VERSION : 1.0
   VAR_INPUT
      IN_iSourceIndex : Int;
      IN_iDestIndex : Int;
      IN_iCount : Int;
   END_VAR
   VAR_IN_OUT
      INO_vSourceArrayStruct : Variant;
      INO_vDestArrayStruct : Variant;
   END_VAR
BEGIN
   #GP_BlockMoveStruct :=  MOVE_BLK_VARIANT(SRC:=#INO_vSourceArrayStruct,
                                            COUNT:=INT_TO_UDINT(#IN_iCount),
                                            SRC_INDEX:=INT_TO_DINT(#IN_iSourceIndex),
                                            DEST_INDEX:=INT_TO_DINT(#IN_iDestIndex),
                                            DEST=>#INO_vDestArrayStruct);
END_FUNCTION

// folder: TaskErrors

ORGANIZATION_BLOCK "Time error interrupt"   // OB80, LAD, TimeErrorInterrupt
{ S7_Optimized_Access := 'TRUE' }
VERSION : 0.1
   VAR_INPUT
      Fault_ID : Byte;   // Fault identifier
      Csg_OBnr : OB_Any;   // Number of OB causing the error
      Csg_Prio : UInt;   // Priority of OB causing the error
   END_VAR
BEGIN
END_ORGANIZATION_BLOCK

ORGANIZATION_BLOCK "Diagnostic error interrupt"   // OB82, LAD, DiagnosticErrorInterrupt
{ S7_Optimized_Access := 'TRUE' }
VERSION : 0.1
   VAR_INPUT
      IO_State : Word;   // IO state of the HW object
      LADDR : Hw_Any;   // Hardware identifier
      Channel : UInt;   // Channel number
      MultiError : Bool;   // =true if more than one error is present
   END_VAR
   VAR_TEMP
      RALM : Struct
         AINFO : "AINFO_";
         TINFO : "TINFO_";
         RETVAL : Int;
         ALLARMI_da_OB82 : Struct
            RALM : "PN_Alarm";
            LADDR : Hw_Any;
            evento_uscente : Bool;
         END_STRUCT;
      END_STRUCT;
      TMP_dId : DInt;
   END_VAR
BEGIN

REGION Network 1
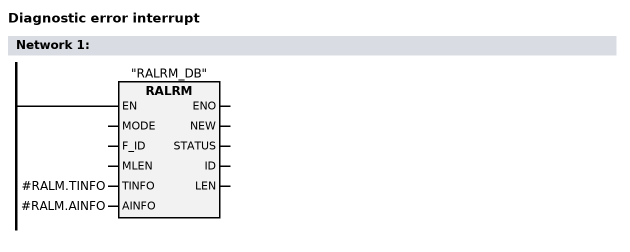
   "RALRM_DB"(TINFO := #RALM.TINFO, AINFO := #RALM.AINFO);   // RALRM
END_REGION

REGION Network 2 (SCL): Set alarms
   #TMP_dId:=UINT_TO_DINT("RALRM_DB".ID);

   IF "RALRM_DB".NEW THEN
       CASE #TMP_dId OF
           1:
               "RALRM_AUX_DB".tAlm.tF.xDevice1 := 1;
           2:
               "RALRM_AUX_DB".tAlm.tF.xDevice2 := 1;
           3:
               "RALRM_AUX_DB".tAlm.tF.xDevice3 := 1;
           4:
               "RALRM_AUX_DB".tAlm.tF.xDevice4 := 1;
           5:
               "RALRM_AUX_DB".tAlm.tF.xDevice5 := 1;
           6:
               "RALRM_AUX_DB".tAlm.tF.xDevice6 := 1;
           7:
               "RALRM_AUX_DB".tAlm.tF.xDevice7 := 1;
           8:
               "RALRM_AUX_DB".tAlm.tF.xDevice8 := 1;
           9:
               "RALRM_AUX_DB".tAlm.tF.xDevice9 := 1;
           10:
               "RALRM_AUX_DB".tAlm.tF.xDevice10 := 1;
           ELSE
               ;
       END_CASE;
   END_IF;
END_REGION
END_ORGANIZATION_BLOCK

ORGANIZATION_BLOCK "Pull or plug of modules"   // OB83, LAD, PullPlug
{ S7_Optimized_Access := 'TRUE' }
VERSION : 0.1
   VAR_INPUT
      LADDR : Hw_Io;   // Hardware identifier
      Event_Class : Byte;   // 16#38/39: module inserted, removed
      Fault_ID : Byte;   // Fault identifier
   END_VAR
BEGIN
END_ORGANIZATION_BLOCK

ORGANIZATION_BLOCK "Rack or station failure"   // OB86, LAD, RackStationFailure
{ S7_Optimized_Access := 'TRUE' }
VERSION : 0.1
   VAR_INPUT
      LADDR : Hw_Device;   // Hardware identifier
      Event_Class : Byte;   // Event class
      Fault_ID : Byte;   // Fault identifier
   END_VAR
BEGIN
END_ORGANIZATION_BLOCK

ORGANIZATION_BLOCK "Programming error"   // OB121, LAD, ProgrammingError
{ S7_Optimized_Access := 'TRUE' }
VERSION : 0.1
   VAR_INPUT
      BlockNr : UInt;   // Number of causing block
      Reaction : USInt;   // 0:ignore, 1:substitute, 2:skip
      Fault_ID : Byte;   // Fault identifier
      BlockType : USInt;   // 16#01:OB, 16#02:FC, 16#03:FB, 16#04:SFC, 16#05:SFB, 16#06:DB: Type of block causing the error
      Area : USInt;   // Area where the error occured
      DBNr : DB_ANY;   // DB number if Area = DB or DI
      Csg_OBNr : OB_Any;   // Number of OB causing the error
      Csg_Prio : USInt;   // Priority of OB causing the error
      Width : USInt;   // 0:bit, 1:byte, 2:word, 3:dword, 4:lword
   END_VAR
BEGIN
END_ORGANIZATION_BLOCK

ORGANIZATION_BLOCK "IO access error"   // OB122, LAD, IOAccessError
{ S7_Optimized_Access := 'TRUE' }
VERSION : 0.1
   VAR_INPUT
      BlockNr : UInt;   // Number of causing block
      Reaction : USInt;   // 0:ignore, 1:substitute, 2:skip
      Fault_ID : Byte;   // 16#42:reading, 16#43:writing
      BlockType : USInt;   // 16#01:OB, 16#02:FC, 16#03:FB, 16#04:SFC, 16#05:SFB, 16#06:DB: Type of block causing the error
      Area : USInt;   // 16#81:I, 16#82:Q: IO area where the IOaccess error occured
      DBNr : DB_ANY;   // Reserved for system
      Csg_OBNr : OB_Any;   // Number of OB causing the error
      Csg_Prio : USInt;   // Priority of OB causing the error
      Width : USInt;   // 0:bit, 1:byte, 2:word, 3:dword, 4:lword
   END_VAR
BEGIN
END_ORGANIZATION_BLOCK

// ===== PLC "1B160AP"  CPU 1512SP-1 PN =====

VAR_GLOBAL   // PLC tag table "Tabella delle variabili standard"
   "System_Byte" AT %MB0 : Byte;
   "FirstScan" AT %M0.0 : Bool;
   "DiagStatusUpdate" AT %M0.1 : Bool;
   "AlwaysTRUE" AT %M0.2 : Bool;
   "AlwaysFALSE" AT %M0.3 : Bool;
   "AlwaysOFF_Debug" AT %M10.0 : Bool;
   "o.1B160AP1.Open_SW_Gate" AT %Q39.0 : Bool;
   "i.1B160AP1.CounterActualValue" AT %ID30 : DWord;
   "i.1B160AP1.FrequencyActualValue" AT %ID38 : Real;
   "i.1B160AP1.CaptureValue" AT %ID34 : DWord;
   "o.1B160AP1.Res_Event" AT %Q40.1 : Bool;
   "o.1B160AP1.M217CutPressureHead1" AT %AW50 : Int;
   "o.1B160AP1.M217CutPressureHead2" AT %AW52 : Int;
   "o.1B160AP1.M217CutPressureHead5" AT %QW58 : Int;
   "o.1B160AP1.Enable_Measure" AT %Q39.7 : Bool;
   "i.1B160AP1.CounterCardStatus" AT %ED42 : DWord;
   "o.1B160AP1.CounterCardStatus" AT %AD38 : DWord;
   "o.1B160AP1.M217CutPressureHead3" AT %AW54 : Int;
   "o.1B160AP1.M217CutPressureHead4" AT %QW56 : Int;
   "o.IDeviceCPU0" AT %Q250.0 : "UDT_CM_IDEV_ToMainLine";
   "i.IDeviceCPU0" AT %I250.0 : "UDT_CM_IDEV_FromMainLine";
   "i.1B160AP1.Res_Event_Ack" AT %I43.1 : Bool;
   "i.1B160AP1.Event_Capture" AT %I45.6 : Bool;
   "cigliu" AT %M1.0 : Bool;
   "i.1B160AP1.1B18-2L+.PowerSupplyInputControlCabinetON" AT %E0.0 : Bool;
   "i.1B160AP1.1B18-3L+.InputInstallationPowerSupplyON" AT %E0.1 : Bool;
   "i.1B160AP1.1B11QF1/2.AnomalyPowerSupplies230V" AT %E0.2 : Bool;
   "i.1B160AP1.1B18QF2.PowerSupply24VLogic" AT %E0.3 : Bool;
   "i.1B160AP1.1B18QF3.PowerSupply24VLogic" AT %E0.4 : Bool;
   "i.1B160AP1.1B20QF2.PowerSupply24VLogic" AT %E0.5 : Bool;
   "i.1B160AP1.1B122KE1.MainEmergencyON" AT %E1.1 : Bool;
   "i.1B160AP1.1B41QF1.ProtectionPowerSupply36V_Motor_1-4" AT %I1.4 : Bool;
   "i.1B160AP1.1B41QF2.ProtectionPowerSupplyMotorsYcut_1-4" AT %I1.5 : Bool;
   "i.1B160AP1.1B51QM1.ProtectionCarriageTranslation" AT %E2.0 : Bool;
   "i.1B160AP1.1B52QM1.ProtectionCarriageTranslation" AT %E2.1 : Bool;
   "i.1B160AP1.1B53QM1.ProtectionCarriageTranslation" AT %E2.2 : Bool;
   "i.1B160AP1.1B54QM1.ProtectionCarriageTranslation" AT %E2.3 : Bool;
   "i.1B160AP1.1B55QM1.ProtectionCarriageTranslation" AT %I2.4 : Bool;
   "i.1B160AP1.M217B1SB1.LocalEmergency" AT %I3.1 : Bool;
   "i.1B160AP1.M217B1SB3_SB4.HeadsUpIstantaneous" AT %I3.0 : Bool;
   "i.1B411AP1.1B411SA1.Head1.CuttingPressure+" AT %E111.2 : Bool;
   "i.1B411AP1.1B411SQ1.Head1.CarriageHeadWorkPosition" AT %E111.3 : Bool;
   "i.1B411AP1.1B411SA1.Head1.CuttingPressure-" AT %E112.2 : Bool;
   "i.1B411AP1.1B411SA2.Head1.ProductionON" AT %E112.4 : Bool;
   "i.1B412AP1.1B412SA1.Head2.CuttingPressure+" AT %E121.2 : Bool;
   "i.1B412AP1.1B412SQ1.Head2.CarriageHeadWorkPosition" AT %E121.3 : Bool;
   "i.1B412AP1.1B412SA1.Head2.CuttingPressure-" AT %E122.2 : Bool;
   "i.1B412AP1.1B412SA2.Head2.ProductionON" AT %E122.4 : Bool;
   "i.1B413AP1.1B413SA1.Head3.CuttingPressure+" AT %E131.2 : Bool;
   "i.1B413AP1.1B413SQ1.Head3.CarriageHeadWorkPosition" AT %E131.3 : Bool;
   "i.1B413AP1.1B413SA1.Head3.CuttingPressure-" AT %E132.2 : Bool;
   "i.1B413AP1.1B413SA2.Head3.ProductionON" AT %E132.4 : Bool;
   "i.1B414AP1.1B414SA1.Head4.CuttingPressure+" AT %E141.2 : Bool;
   "i.1B414AP1.1B414SQ1.Head4.CarriageHeadWorkPosition" AT %E141.3 : Bool;
   "i.1B414AP1.1B414SA1.Head4.CuttingPressure-" AT %E142.2 : Bool;
   "i.1B414AP1.1B414SA2.Head4.ProductionON" AT %E142.4 : Bool;
   "i.1B415AP1.1B415SA1.Head5.CuttingPressure+" AT %I151.2 : Bool;
   "i.1B415AP1.1B415SQ1.Head5.CarriageHeadWorkPosition" AT %I151.3 : Bool;
   "i.1B415AP1.1B415SA1.Head5.CuttingPressure-" AT %I152.2 : Bool;
   "i.1B415AP1.1B415SA2.Head5.ProductionON" AT %I152.4 : Bool;
   "o.1B160AP1.1B251HL1.AreaFailure" AT %A0.0 : Bool;
   "o.1B160AP1.1B251KA1.ResetLocalEmergency" AT %A0.2 : Bool;
   "o.1B160AP1.EnableCard1" AT %A2.0 : Bool;
   "o.1B160AP1.EnableCard2" AT %A2.1 : Bool;
   "o.1B160AP1.EnableCard3" AT %A2.2 : Bool;
   "o.1B160AP1.EnableCard4" AT %A2.3 : Bool;
   "o.1B160AP1.EnableCard5" AT %Q2.4 : Bool;
   "o.1B160AP1.M217B1HL5.MachineToMaintenance" AT %Q0.6 : Bool;
   "o.1B160AP1.M217B1HL3.MachineReady" AT %Q0.4 : Bool;
   "o.1B160AP1.M217B1HL6.MachineOutOfOrder" AT %Q0.7 : Bool;
   "o.1B160AP1.M217B1HL4.MachineInOrder" AT %Q0.5 : Bool;
   "o.1B411AP1.1B411YV2.Head1.CuttingLubrication" AT %A111.0 : Bool;
   "o.1B411AP1.1B411YV1.Head1.CuttingHeadGlassApproach" AT %A111.1 : Bool;
   "o.1B411AP1.1B411SA2.Head1.ProductionON" AT %A111.4 : Bool;
   "o.1B412AP1.1B412YV2.Head2.CuttingLubrication" AT %A121.0 : Bool;
   "o.1B412AP1.1B412YV1.Head2.CuttingHeadGlassApproach" AT %A121.1 : Bool;
   "o.1B412AP1.1B412SA2.Head2.ProductionON" AT %A121.4 : Bool;
   "o.1B413AP1.1B413YV2.Head3.CuttingLubrication" AT %A131.0 : Bool;
   "o.1B413AP1.1B413YV1.Head3.CuttingHeadGlassApproach" AT %A131.1 : Bool;
   "o.1B413AP1.1B413SA2.Head3.ProductionON" AT %A131.4 : Bool;
   "o.1B414AP1.1B414YV2.Head4.CuttingLubrication" AT %A141.0 : Bool;
   "o.1B414AP1.1B414YV1.Head4.CuttingHeadGlassApproach" AT %A141.1 : Bool;
   "o.1B414AP1.1B414SA2.Head4.ProductionON" AT %A141.4 : Bool;
   "o.1B415AP1.1B415YV2.Head5.CuttingLubrication" AT %Q151.0 : Bool;
   "o.1B415AP1.1B415YV1.Head5.CuttingHeadGlassApproach" AT %Q151.1 : Bool;
   "o.1B415AP1.1B415SA2.Head5.ProductionON" AT %Q151.4 : Bool;
   "i.1B160AP1.1B20QF3.PowerSupply24VLogic" AT %I0.6 : Bool;
   "i.1B160AP1.1B42QF1.ProtectionPowerSupply36V_Motor_5-8" AT %I1.6 : Bool;
   "i.1B160AP1.1B42QF2.ProtectionPowerSupplyMotorsYcut_5-8" AT %I1.7 : Bool;
   "i.1B160AP1.1B56QM1.ProtectionCarriageTranslation" AT %I2.5 : Bool;
   "i.1B160AP1.1B57QM1.ProtectionCarriageTranslation" AT %I2.6 : Bool;
   "i.1B160AP1.1B58QM1.ProtectionCarriageTranslation" AT %I2.7 : Bool;
   "o.1B160AP1.EnableCard6" AT %Q2.5 : Bool;
   "o.1B160AP1.EnableCard7" AT %Q2.6 : Bool;
   "o.1B160AP1.EnableCard8" AT %Q2.7 : Bool;
   "o.1B160AP1.M217CutPressureHead6" AT %QW60 : Int;
   "o.1B160AP1.M217CutPressureHead7" AT %QW62 : Int;
   "o.1B160AP1.M217CutPressureHead8" AT %QW64 : Int;
   "o.1B416AP1.1B416SA2.Head6.ProductionON" AT %Q161.4 : Bool;
   "o.1B416AP1.1B416YV1.Head6.CuttingHeadGlassApproach" AT %Q161.1 : Bool;
   "o.1B416AP1.1B416YV2.Head6.CuttingLubrication" AT %Q161.0 : Bool;
   "o.1B417AP1.1B417SA2.Head7.ProductionON" AT %Q171.4 : Bool;
   "o.1B417AP1.1B417YV1.Head7.CuttingHeadGlassApproach" AT %Q171.1 : Bool;
   "o.1B417AP1.1B417YV2.Head7.CuttingLubrication" AT %Q171.0 : Bool;
   "o.1B418AP1.1B418SA2.Head8.ProductionON" AT %Q181.4 : Bool;
   "o.1B418AP1.1B418YV1.Head8.CuttingHeadGlassApproach" AT %Q181.1 : Bool;
   "o.1B418AP1.1B418YV2.Head8.CuttingLubrication" AT %Q181.0 : Bool;
   "i.1B416AP1.1B416SA1.Head6.CuttingPressure-" AT %I162.2 : Bool;
   "i.1B416AP1.1B416SA1.Head6.CuttingPressure+" AT %I161.2 : Bool;
   "i.1B416AP1.1B416SA2.Head6.ProductionON" AT %I162.4 : Bool;
   "i.1B416AP1.1B416SQ1.Head6.CarriageHeadWorkPosition" AT %I161.3 : Bool;
   "i.1B417AP1.1B417SA1.Head7.CuttingPressure-" AT %I172.2 : Bool;
   "i.1B417AP1.1B417SA1.Head7.CuttingPressure+" AT %I171.2 : Bool;
   "i.1B417AP1.1B417SA2.Head7.ProductionON" AT %I172.4 : Bool;
   "i.1B417AP1.1B417SQ1.Head7.CarriageHeadWorkPosition" AT %I171.3 : Bool;
   "i.1B418AP1.1B418SA1.Head8.CuttingPressure-" AT %I182.2 : Bool;
   "i.1B418AP1.1B418SA1.Head8.CuttingPressure+" AT %I181.2 : Bool;
   "i.1B418AP1.1B418SA2.Head8.ProductionON" AT %I182.4 : Bool;
   "i.1B418AP1.1B418SQ1.Head8.CarriageHeadWorkPosition" AT %I181.3 : Bool;
   "i.1B160AP1.M217B1SB2.LocalEmergency" AT %I3.2 : Bool;
END_VAR

VAR_GLOBAL CONSTANT   // PLC tag table "Tabella delle variabili standard"
   "CONST_dNumberOfHeadsCycle" : DInt := 7;   // Number of heads / Number of heads-1
   "CONST_dNumberOfHeads" : DInt := 8;   // Number of heads-1 / Number of heads
   "CONST_dPressureMax_MN" : DInt := 180000;   // Maximum allowable pressure [N/1000]
   "CONST_dPressureMin_MN" : DInt := 0;   // Minimum allowable pressure [N/1000]
   "CONST_dPressureMax_Unit" : DInt := 27648;   // Maximum allowable pressure Analog unit
   "CONST_dPressureMin_Unit" : DInt := 0;   // Minimum allowable pressure Analog unit
   "CONST_dFire_OnOff_MaxValue" : DInt := 5000;   // Fire ON OFF max value [mm/100]
   "CONST_dFire_OnOff_MinValue" : DInt := 0;   // Fire ON OFF min value [mm/100]
   "CONST_dPressureMax_Display_MN" : DInt := 180000;   // Maximum allowable pressure [N/1000]
   "CONST_dPressureMin_Display_MN" : DInt := 0;   // Minimum allowable pressure [N/1000]
   "CONST_dPressureMax_Display_Unit" : DInt := 27648;   // Maximum allowable pressure Analog unit
   "CONST_dPressureMin_Display_Unit" : DInt := 0;   // Minimum allowable pressure Analog unit
   "CONST_dPressureIncreasePneumatic_MN" : DInt := 250000;   // Pressure increse by cylinder [N/1000]
END_VAR

TYPE "ILx2T_Ref"
AUTHOR : SEMotion
FAMILY : LXM32
VERSION : 0.5
   STRUCT
      i_woDriveStatus : Word;
      i_by_ModeStatus : Byte;
      i_by_driveInput : Byte;
      i_wo_ActionWord : Word;
      i_wo_SpecialFunctions : Word;
      q_wo_dmControl : Word;
      q_dw_refA_16 : Word;
      q_dw_refB_32 : DWord;
      arOutputData : Array[0..7] of Byte;
      arInputData : Array[0..7] of Byte;
      stDriveStatus : Struct
         HaltActive : Bool;   // HALT is active
         reserved_Bit9 : Bool;
         reserved_Bit10 : Bool;
         reserved_Bit11 : Bool;
         reserved_Bit12 : Bool;
         x_Add : Bool;   // additional information
         x_End : Bool;   // OP mode finished - standstill
         x_Err : Bool;   // error
         state_Bit0 : Bool;   // Drive state bit 0
         state_Bit1 : Bool;   // Drive state bit 1
         state_Bit2 : Bool;   // Drive state bit 2
         state_Bit3 : Bool;   // Drive state bit 3
         reseverd_Bit4 : Bool;
         reserved_Bit5 : Bool;
         FaultActive : Bool;   // FAULT is active
         WarningActive : Bool;   // WARNING is active
      END_STRUCT;
      st_ModeStatus : Struct
         Mode_0 : Bool;   // Actual OP mode bit 0
         Mode_1 : Bool;   // Actual OP mode bit 1
         Mode_2 : Bool;   // Actual OP mode bit 2
         Mode_3 : Bool;   // Actual OP mode bit 3
         reserved : Bool;
         Reference_OK : Bool;   // drive is referenced
         ModeError : Bool;   // Status mode error
         ModeToggle : Bool;   // Status mode toggle
      END_STRUCT;
      st_ActionWord : Struct
         MotionNegative : Bool;   // negative direction
         InsidePosWindow : Bool;   // Inside Position Window
         reserved_Bit10 : Bool;
         TargetVelocityZero : Bool;   // Target velocity is zero
         Decelerating : Bool;
         Accelerating : Bool;
         ConstantVelocity : Bool;
         reserved_Bit15 : Bool;
         Reserved : Bool;
         Reserved_1 : Bool;
         Reserved_2 : Bool;
         Reserved_3 : Bool;
         Reserved_4 : Bool;
         Reserved_5 : Bool;
         MotionZero : Bool;   // Motion zero, actual velocity is zero
         MotionPositive : Bool;   // motor is moving in positiove direction
      END_STRUCT;
      st_SpecFunctions : Struct
         reserved_4 : Bool;   // Capture counter channel 1 bit 0
         reserved_5 : Bool;   // Capture counter channel 1 bit 1
         reserved_6 : Bool;   // Capture counter channel 2 bit 0
         reserved_7 : Bool;   // Capture counter channel 2 bit 1
         reserved_12 : Bool;
         reserved_13 : Bool;
         reserved_14 : Bool;
         reserved_15 : Bool;
         CAP1_0 : Bool;   // Actual OP mode bit 0
         CAP1_1 : Bool;   // Actual OP mode bit 1
         CAP2_0 : Bool;   // Actual OP mode bit 2
         CAP2_1 : Bool;   // Actual OP mode bit 3
         reserved : Bool;   // Actual OP mode bit 4
         reserved_1 : Bool;   // Status ModeDataError
         reserved_2 : Bool;   // Status mode error
         reserved_3 : Bool;   // Status mode toggle
      END_STRUCT;
      InitAccessID : Int;   // AccessID counter for INIT
      ProChAccessID : Int;   // Access ID Processchannel
      ParChAccessID : Int;   // Access ID Parameterchannel
      x_QuickStopInt : Bool;   // Library internal QuickStop Command
      x_FaultResetInt : Bool;   // Library internal FaultReset Command
      x_Set_HALT_Int : Bool;   // Library internal Set HALT Command
      x_Clear_HALT_Int : Bool;   // Library internal Clear HALT Command
      x_Continue_Int : Bool;   // Library internal HALT Contimue Command
      by_OP_ModeAct : Byte;   // Status - Actual operation mode
      x_IO_1 : Bool;   // Status of digital IO 1 (Bit 0)
      x_IO_2 : Bool;   // Status of digital IO 2 (Bit 1)
      x_IO_3 : Bool;   // Status of digital IO 3 (Bit 2)
      x_IO_4 : Bool;   // Status of digital IO 4 (Bit 3)
      x_STO_A : Bool;   // Status of Safe Torque Off Channel A
      x_STO_B : Bool;   // Status of Safe Torque Off Channel B
      x_reserved_6 : Bool;
      x_reserved_7 : Bool;
      x_CommandWriteParameter : Bool;
      x_CommandReadParameter : Bool;
      x_StatusReadParameter_OK : Bool;
      x_StatusReadParameter_Error : Bool;
      x_Status_WriteParameter_OK : Bool;
      x_Status_WriteParameter_Error : Bool;
      di_ParameterReadValue : DInt;
      di_ParameterWriteValue : DInt;
      udi_ModbusAddress_Read : UDInt;
      udi_ModbusAddress_Write : UDInt;
   END_STRUCT;
END_TYPE

TYPE "UDT_DataManager_HeadsBuffer"
VERSION : 0.1
   STRUCT
      rgdMissionID : Array[0..20] of DInt;   // Head#x mission ID
      rgdRequestPosition_cmm : Array[0..20] of DInt;   // Head#x request position [mm/100]
      rgdFireRequest : Array[0..20] of DInt;   // Head#x fire request
      dNumberOfElement : DInt;   // Number of element inside the buffer
   END_STRUCT;
END_TYPE

TYPE "UDT_DataManager_Insert"
VERSION : 0.1
   STRUCT
      dMissionCode : DInt;   // Mission code
      dMissionStart_cmm : DInt;   // Mission counter start [mm/100]
      dMissionEnd_cmm : DInt;   // Mission counter end [mm/100]
      rgxFireRequest : Array[0.."CONST_dNumberOfHeadsCycle"] of Bool;   // Fire request missions
      rgdHeadsPosition_cmm : Array[0.."CONST_dNumberOfHeadsCycle"] of DInt;   // Head#x position request [mm/100]
      xNewMission : Bool;   // New mission available
      xSystemReset : Bool;   // System reset
      rgdArmONReaction_ms : Array[0.."CONST_dNumberOfHeadsCycle"] of DInt;   // Head#x arm ON reaction [ms]
      rgdArmOFFReaction_ms : Array[0.."CONST_dNumberOfHeadsCycle"] of DInt;   // Head#x arm OFF reaction [ms]
      rgdFireONReaction_ms : Array[0.."CONST_dNumberOfHeadsCycle"] of DInt;   // Head#x fire ON reaction [ms]
      rgdFireOFFReaction_ms : Array[0.."CONST_dNumberOfHeadsCycle"] of DInt;   // Head#x fire OFF reaction [ms]
      rgdOilDelayStart_ms : Array[0.."CONST_dNumberOfHeadsCycle"] of DInt;   // Head#x oil delay start [ms]
      rgdOilDelayEnd_ms : Array[0.."CONST_dNumberOfHeadsCycle"] of DInt;   // Head#x oil advance end [ms]
      rgdFireONDelayStart_cmm : Array[0.."CONST_dNumberOfHeadsCycle"] of DInt;   // Head#x fire ON delay start [mm/100]
      rgdFireOFFDelayEnd_cmm : Array[0.."CONST_dNumberOfHeadsCycle"] of DInt;   // Head#x fire OFF delay end [mm/100]
   END_STRUCT;
END_TYPE

TYPE "UDT_DataManager"
VERSION : 0.1
   STRUCT
      tInputData : "UDT_DataManager_Insert";   // Manager input data
      tOutputData : "UDT_DataManager_Output";   // Manager output data
      dInterruptNumMissionTank : DInt;   // Number of mission fire inside the tank
      rgtInterruptMissionTank : Array[0..20] of "UDT_DataManager_Tank";   // Array of fire missions
      rgtOilList : Array[0.."CONST_dNumberOfHeadsCycle"] of "UDT_DataManager_HeadsBuffer";   // Oil list manager
      rgtArmList : Array[0.."CONST_dNumberOfHeadsCycle"] of "UDT_DataManager_HeadsBuffer";   // Arm list manager
   END_STRUCT;
END_TYPE

TYPE "UDT_DataManager_Output"
VERSION : 0.1
   STRUCT
      dMissionCode : DInt;   // Mission code number
      rgdFireHeadThreshold_cmm : Array[0.."CONST_dNumberOfHeadsCycle"] of DInt;   // Head#x firing threshold [mm/100]
      rgdHeadsPositions_cmm : Array[0.."CONST_dNumberOfHeadsCycle"] of DInt;   // Head#x positions request [mm/100]
      rgxFireHeadON_OFF : Array[0.."CONST_dNumberOfHeadsCycle"] of Bool;   // Head#x firing type request [bit]
      rgxDataToProcessInter : Array[0.."CONST_dNumberOfHeadsCycle"] of Bool;   // Head#x data to process by interrupt
      xGateOpen : Bool;   // Interrupt gate open
      dTargetLineValue_cmm : DInt;   // Virtual target line value [mm/100]
      rgxArmRequest : Array[0.."CONST_dNumberOfHeadsCycle"] of Bool;   // Head#x arming request
      rgdArmRequestTarget_cmm : Array[0.."CONST_dNumberOfHeadsCycle"] of DInt;   // Arm request target virtual [mm/100]
      rgxOilRequest : Array[0.."CONST_dNumberOfHeadsCycle"] of Bool;   // Head#x oil request
      rgdOilRequestTarget_cmm : Array[0.."CONST_dNumberOfHeadsCycle"] of DInt;   // Oil request target virtual [mm/100]
      rgdArmRequestIDMission : Array[0.."CONST_dNumberOfHeadsCycle"] of DInt;   // Arm request ID mission
      rgdOilRequestIDMission : Array[0.."CONST_dNumberOfHeadsCycle"] of DInt;   // Oil request ID mission
   END_STRUCT;
END_TYPE

TYPE "UDT_DataManager_Tank"
VERSION : 0.1
   STRUCT
      dMissionCode : DInt;   // Mission code
      dMissionValue_cmm : DInt;   // Mission value [mm/100]
      rgxFireRequest : Array[0.."CONST_dNumberOfHeadsCycle"] of Bool;   // Head#x fire request
      rgdHeadsPositions_cmm : Array[0.."CONST_dNumberOfHeadsCycle"] of DInt;   // Head#x position request [mm/100]
   END_STRUCT;
END_TYPE

TYPE "UDT_MB_ConnData"
   STRUCT
      IP_OCTET_1 : USInt;
      IP_OCTET_2 : USInt;
      IP_OCTET_3 : USInt;
      IP_OCTET_4 : USInt;
      ConnectID1 : Conn_Ouc;
      ConnectID2 : Conn_Ouc;
      ConnectID3 : Conn_Ouc;
      ConnectID4 : Conn_Ouc;
   END_STRUCT;
END_TYPE

TYPE "UDT_CM_IDEV_FromMainLine"
VERSION : 0.1
   STRUCT
      dSpare1 : Array[0..2] of DInt;
      xCycleON : Bool;   // Cycle ON
      xResetAnomaly : Bool;   // Reset anomaly
      xResetBuffers : Bool;   // Reset buffer
      xGlassBreak : Bool;   // Glass break under the bridge
      xPLCActive0 : Bool;   // PLC Active (0=CPU0, 1=CPU1)
      xPLCActive1 : Bool;   // PLC Active (0=CPU0, 1=CPU1)
      xQLTplate : Bool;   // Quality plate in progress
      xSpare2 : Bool;
      xSpare3 : Bool;
      xSpare4 : Bool;
      xSpare5 : Bool;
      xSpare6 : Bool;
      xSpare7 : Bool;
      xSpare8 : Bool;
      xSpare9 : Bool;
      xSpare10 : Bool;
      xStatusSpare : Array[0..15] of Bool;
      dSpare2 : Array[0..7] of DInt;
      iSpare : Int;
   END_STRUCT;
END_TYPE

TYPE "UDT_CM_IDEV_ToMainLine"
VERSION : 0.1
   STRUCT
      dProcessingIDPlate : DInt;   // Processing ID Plate [Num]
      dSpare1 : DInt;
      dSpare2 : DInt;
      rgxStatus : Array[0..31] of Bool;   // Status heads
      rgdHeadsPositions_cmm : Array[0..15] of DInt;   // Head #x position status
      rgxHeadStatus : Array[0..15] of Bool;   // Head #x enabled
      rgxCuttingStatus : Array[0..15] of Bool;   // Head #x cuuting status
      rgdHeadsPressure : Array[0..15] of DInt;   // Head #x Pressure [mN]
      rgrHeadsSpace : Array[0..15] of Real;   // Head #x Distance [Km]
      iFireOffset_ON : Int;   // All head fire on offset
      iFireOffset_OFF : Int;   // All head fire off offset
      iSpare : Int;
      dSpare : Array[0..7] of DInt;
   END_STRUCT;
   // // rgxStatus[0] : Glass break in progress
   // // rgxStatus[1] : Liftup pushbutton engaged
   // // rgxStatus[2] : Bridge enabled
   // // rgxStatus[3] : Bridge locked
   // // rgxStatus[8] : Fire offset calibration
END_TYPE

TYPE "UDT_CM_RECV_SyncroData"
VERSION : 0.1
   STRUCT
      dMissionID : DInt;   // Mission Identifier
      dSynchroValue_cmm : DInt;   // Counter value in the last synchro [mm/100]
      dSpare : Array[0..7] of DInt;
      xSpare : Array[0..15] of Bool;
      dSpare2 : Array[0..2] of DInt;
      iSpare : Int;
   END_STRUCT;
END_TYPE

TYPE "UDT_CM_RECV_MissionData"
VERSION : 0.1
   STRUCT
      dMissionID : DInt;   // Mission Identifier
      dMissionStart_cmm : DInt;   // Mission counter start [mm/100]
      dMissionEnd_cmm : DInt;   // Mission counter stop [mm/100]
      dTrackingDbNumber : DInt;   // Tracking DB number
      dSpare1 : Array[0..9] of DInt;
      rgxFireRequest : Array[0..31] of Bool;   // Head #x firing request
      rgdHeadsPosition_cmm : Array[0..15] of DInt;   // Head #x position request [mm/100]
      dSpare2 : Array[0..14] of DInt;
   END_STRUCT;
END_TYPE

TYPE "UDT_CM_Manager"
VERSION : 0.1
   STRUCT
      ST_xNewDataReceiveCPU0 : Bool;   // New data receive
      ST_xErrorCPU0 : Bool;   // Error
      ST_xNewSynchCPU0 : Bool;   // New synch
      ST_xNewMissionCPU0 : Bool;   // New mission
      AUX_iDataLenghtCPU0 : Word;   // Data lenght
      AUX_iStateCPU0 : Int;   // Status
      ST_xNewDataReceiveCPU1 : Bool;   // New data receive
      ST_xErrorCPU1 : Bool;   // Error
      ST_xNewSynchCPU1 : Bool;   // New synch
      ST_xNewMissionCPU1 : Bool;   // New mission
      AUX_iDataLenghtCPU1 : Word;   // Data lenght
      AUX_iStateCPU1 : Int;   // Status
      AUX_tmON_ConsumedTimeout : IEC_TIMER;   // Timer ON consumed timeout PLCA
      AUX_rgdHeadMissionIDInProg_Copy : Array[0.."CONST_dNumberOfHeadsCycle"] of DInt;   // Head#x mission ID in progress
      AUX_rgxHeadFiringMissionInProg_Copy : Array[0.."CONST_dNumberOfHeadsCycle"] of Bool;   // Head#x firing mission in progress
      ST_xConsumedTimeout : Bool;   // Consumed message timeout PLCA
      ST_xMissionPacketLost : Bool;   // Mission message packet lost PLC A
      ST_xSyncroPacketLost : Bool;   // Syncro message packet lost PLC A
      ST_MutingFiringOB : Bool;   // Muting Ob30 firing
   END_STRUCT;
END_TYPE

TYPE "UDT_HeadPar"
VERSION : 0.1
   STRUCT
      iAddress : Int;
      iLength : Byte;
      dValue : DInt;
   END_STRUCT;
END_TYPE

TYPE "UDT_AxisParameters"
VERSION : 0.1
   STRUCT
      rgtAxisParameters : Array[0..20] of "UDT_HeadPar";
      dParametersToDownload : DInt;
   END_STRUCT;
END_TYPE

TYPE "UDT_BRCV_FromMainLine"
VERSION : 0.1
   STRUCT
      SyncroData : "UDT_CM_RECV_SyncroData";
      MissionData : "UDT_CM_RECV_MissionData";
   END_STRUCT;
END_TYPE

TYPE "LPD_typeCountFeedbackCh"
VERSION : 0.1
   STRUCT
      countValue : DInt := 16#0000;   // Current count value
      capturedValue : DInt := 16#0000;   // Last Capture value acquired
      measuredValue : Real := 0.0;   // Current measured value
      powerError : Bool := FALSE;   // Incorrect supply voltage L+
      encError : Bool := FALSE;   // Incorrect encoder signal
      ldError : Bool := FALSE;   // Error when loading via control interface
      reserved1 : Bool := FALSE;   // Reserved
      reserved2 : Bool := FALSE;   // Reserved
      reserved3 : Bool := FALSE;   // Reserved
      reserved4 : Bool := FALSE;   // Reserved
      reserved5 : Bool := FALSE;   // Reserved
      commActive : Bool := FALSE;   // Comm active
      resEventAck : Bool := FALSE;   // Reset of event bits active
      ldStsSlot0 : Bool := FALSE;   // Load request for Slot 0 detected and executed (toggling)
      ldStsSlot1 : Bool := FALSE;   // Load request for Slot 1 detected and executed (toggling)
      stsReady : Bool := FALSE;   // Digital on-board I/O started up and parameters assigned
      stsSwGate : Bool := FALSE;   // Software gate status
      reserved7 : Bool := FALSE;   // Reserved
      reserved8 : Bool := FALSE;   // Reserved
      stsDir : Bool := FALSE;   // Direction of last count value change
      stsCount : Bool := FALSE;   // Count pulse detected within last approx. 0.5 s
      stsGate : Bool := FALSE;   // Internal gate status
      stsDQ0 : Bool := FALSE;   // Status HSC DQ0
      stsDQ1 : Bool := FALSE;   // Status HSC DQ1
      stsDI0 : Bool := FALSE;   // Status HSC DI0
      stsDI1 : Bool := FALSE;   // Status HSC DI1
      stsDI2 : Bool := FALSE;   // Status HSC DI2
      eventZero : Bool := FALSE;   // Zero crossing has occurred
      eventUnderflow : Bool := FALSE;   // Underflow has occurred
      eventOverflow : Bool := FALSE;   // Overflow has occurred
      eventCompare0 : Bool := FALSE;   // Comparison event for DQ0 has occurred
      eventCompare1 : Bool := FALSE;   // Comparison event for DQ1 has occurred
      eventSync : Bool := FALSE;   // Synchronization has occurred
      eventCapture : Bool := FALSE;   // Capture event has occurred
      stsMeasInterval : Bool := FALSE;   // Count pulse detected in previous measuring interval
   END_STRUCT;
END_TYPE

TYPE "LPD_typeCountControlCh"
VERSION : 0.1
   STRUCT
      loadValue0 : DWord := 16#0000;   // Load value 0
      loadValue1 : DWord := 16#0000;   // Load value 1
      controlByte : Byte := B#16#00;   // Control byte load value
      swGate : Bool := FALSE;   // Software gate
      tmCtrlDQ0 : Bool := FALSE;   // Enable technological function DQ0
      tmCtrlDQ1 : Bool := FALSE;   // Enable technological function DQ1
      setDQ0 : Bool := FALSE;   // Set DQ0
      setDQ1 : Bool := FALSE;   // Set DQ1
      enSyncUp : Bool := FALSE;   // Enable upward synchronization
      enSyncDown : Bool := FALSE;   // Enable downward synchronization
      enCapture : Bool := FALSE;   // Enable capture function
      resError : Bool := FALSE;   // Reset of saved error states
      resEvent : Bool := FALSE;   // Reset of saved events
      reserved0 : Bool := FALSE;   // Reserved
      reserved1 : Bool := FALSE;   // Reserved
      reserved2 : Bool := FALSE;   // Reserved
      reserved3 : Bool := FALSE;   // Reserved
      reserved4 : Bool := FALSE;   // Reserved
      SetDir : Bool := FALSE;   // Count direction (with encoder without direction signal)
      reserved5 : Byte;   // Reserved
   END_STRUCT;
END_TYPE

// folder: ProfinetDiagnostic

TYPE "TINFO_"
VERSION : 0.1
   STRUCT
      OB_start_info : Array[0..19] of Byte;
      W_20_STATION : Word;
      B22_slave_type : Byte;
      B23_interrupt_type : Byte;
      B24_origination : Byte;
      B25_diag_flag : Byte;
      W26_PN_ID : Word;
      W28_MFG_ID : Word;
      W30_INST_ID : Word;
      other_data : Array[1..70] of Byte;
   END_STRUCT;
END_TYPE

TYPE "AINFO_"
VERSION : 0.1
   STRUCT
      W0_block_type : Word;
      W2_block_length : Word;
      W4_version : Word;
      W6_interrupt_type : Word;
      D8_API : DWord;
      W12_comp_slot_num : Word;
      W14_submodule_slot_num : Word;
      D16_module_ID : DWord;
      D20_submodule_ID : DWord;
      W24_interrupt_specifer : Word;
      Add_W0_format_ID : Word;
      Add_W2_channel_num : Word;
      Add_B4_error_info : Byte;
      Add_B5_data_format : Byte;
      Add_W6_error_type : Word;
      extended_info : Array[34..1431] of Byte;
   END_STRUCT;
END_TYPE

TYPE "PN_Alarm"
VERSION : 0.1
   STRUCT
      word_allarme : Word;
      canale : Int;
   END_STRUCT;
END_TYPE

// folder: (top level)

DATA_BLOCK "PLANT_CONSTANTS"   // DB6
{ S7_Optimized_Access := 'TRUE' }
VERSION : 0.1
   VAR
      CONST_rgxHomeSide : Array[0.."CONST_dNumberOfHeadsCycle"] of Bool;   // Head#x home side [0=Operator Side 1=Opposite operator side]
      CONST_dHOpSideEnc_cmm : Array[0.."CONST_dNumberOfHeadsCycle"] of DInt;   // Operator side head encumbrance [mm/100]
      CONST_dHOppoSideEnc_cmm : Array[0.."CONST_dNumberOfHeadsCycle"] of DInt;   // Opposite operatore side encumbrance [mm/100]
      CONST_rgtHeadPar : Array[0.."CONST_dNumberOfHeadsCycle"] of "UDT_AxisParameters";   // Array of head parameters
   END_VAR
BEGIN
   CONST_rgxHomeSide[0] := false;
   CONST_rgxHomeSide[1] := false;
   CONST_rgxHomeSide[2] := true;
   CONST_rgxHomeSide[3] := true;
END_DATA_BLOCK

DATA_BLOCK "M256_Manag_IDB"   // DB7
{ S7_Optimized_Access := 'TRUE' }
VERSION : 0.1
// stored: InstanceOfName M256_Manager
"M256_Manager"
BEGIN
   M256A_IDB[0].tHMW.dDescentReactTime_ms := 2000;
   M256A_IDB[0].tHMW.dRaiseReactTime_ms := -100;
END_DATA_BLOCK

DATA_BLOCK "Z256_Manager"   // DB9
{ S7_Optimized_Access := 'TRUE' }
VERSION : 0.1
BEGIN
END_DATA_BLOCK

DATA_BLOCK "Z256"   // DB13
{ S7_Optimized_Access := 'TRUE' }
VERSION : 0.1
   VAR
      tmOFF_ResetAlarm : IEC_TIMER;   // Reset alarm
      tmON_24Vdc : IEC_TIMER;   // Presence 24Vdc timer
      tmON_EmergencyOK : IEC_TIMER;   // Emergency OK timer
      ST_xZoneError : Bool;   // Zone error
      ST_xSelectionAutoMode : Bool;   // Automatic mode selection
      ST_xSelectionManualMode : Bool;   // Manual mode selection
      ST_xConditionOKManualMode : Bool;   // Condition OK for manual mode
      ST_xManualModeAccepted : Bool;   // Manual mode accepted
      ST_xAutoModeAccepted : Bool;   // Automatic mode accepted
      ST_xManualModeRequest : Bool;   // Manual mode request
      ST_xFaultsEnabled : Bool;   // Faults enabled
      ST_xZoneEmergency : Bool;   // Cumulative of emergency faults active
      ST_xZoneFaults : Bool;   // Cumulative of zone faults
      ST_xZoneStoppingFaults : Bool;   // Cumulative of zone stopping faults
      ST_xZoneWarnings : Bool;   // Cumulative of zone warning
      ST_xGlassBreak : Bool;   // Glass break under the zone
      ST_xConditionOkBridgeOutProd : Bool;   // Condition OK for bridge out of production
      ST_rgxConditionOkHeadOutProd : Array[0.."CONST_dNumberOfHeadsCycle"] of Bool;   // Condition OK for head out of production
      ST_xCycleON : Bool;   // Zone in cycle ON
      ST_xPLCB_Active : Bool;   // PLC B is active
      OSN_xGateOpen : Bool;   // OSN gate open
      OSR_xGateOpen : Bool;   // OSR gate open
      OS_xGeneralReset : Bool;   // General reset
      OS_xGateOpen : Bool;   // OS gate open
      ON_xGateOpen : Bool;   // ON gate open
      INPUT_xOperatorOverstroke : Bool;   // Operator side head overstroke
      INPUT_xOppoOperatorOverstroke : Bool;   // Opposite operator side head overstroke
      INPUT_xInputCtrlCabinetON : Bool;   // L+.Power supply input control cabinet ON
      INPUT_xInputPowerSupplyON : Bool;   // L+.Input installation power supply ON
      INPUT_xAnomalyPower120_240 : Bool;   // QF.Anomaly power supplies 120 / 240
      INPUT_xPowerSupply24vLogic1 : Bool;   // QF.Power supply 24v logic #1
      INPUT_xPowerSupply24vLogic2 : Bool;   // QF.Power supply 24v logic #2
      INPUT_xPowerSupply24vLogic3 : Bool;   // QF.Power supply 24v logic #3
      INPUT_xPowerSupply24vLogic4 : Bool;   // QF.Power supply 24v logic #4
      INPUT_xPowerSupply24vLogic5 : Bool;   // QF.Power supply 24v logic #5
      INPUT_xLocalEmergencyON : Bool;   // KE.Main emergency ON
      INPUT_xMainEmergencyON : Bool;   // KE.Main emergency ON
      INPUT_xProtSupply36v_1 : Bool;   // QF.Protection power supply 36v #1
      INPUT_xProtSupply36v_2 : Bool;   // QF.Protection power supply motors longitudinal cutting #1
      INPUT_xProtMotorLC_1 : Bool;   // QF.Protection power supply 36v #2
      INPUT_xProtMotorLC_2 : Bool;   // QF.Protection power supply motors longitudinal cutting #2
      INPUT_xProtConditioners : Bool;   // QF.Protection conditioners
      INPUT_xResetLocalEmergency : Bool;   // SB.Reset local emergency
      INPUT_xLocalEmergency_SB1 : Bool;   // SB1.Local emergency
      INPUT_xLocalEmergency_SB2 : Bool;   // SB2.Local emergency
      INPUT_xLocalEmergency_Cabinet : Bool;   // Cabinet.Local emergency
      INPUT_rgxHeadsInProduction : Array[0.."CONST_dNumberOfHeadsCycle"] of Bool;   // SL.Head#x in production
      OUTPUT_xResetLocalEmergency : Bool;   // KM.Reset local emergency
      OUTPUT_xAreaFailure : Bool;   // HL.Cabinet area failure
      OUTPUT_xLocalEmergencyON : Bool;   // HL.Local emergency ON
      OUTPUT_xMachineOutOfOrder : Bool;   // HL.Machine out of order RED
      OUTPUT_xMachineToMaintenance : Bool;   // HL.Machine to maintenance YELLOW
      OUTPUT_xMachineInOrder : Bool;   // HL.Machine in order GREEN
      OUTPUT_xMachineReady : Bool;   // HL.Machine ready WHITE
      OUTPUT_rgxHeadsInProduction : Array[0.."CONST_dNumberOfHeadsCycle"] of Bool;   // HL.Head #x in production
   END_VAR
BEGIN
END_DATA_BLOCK

DATA_BLOCK "Z256_hmi"   // DB14
{ S7_Optimized_Access := 'TRUE' }
VERSION : 0.1
   VAR RETAIN
      tHMR : Struct   // {[Unit][Scada unit][Low limit][High limit][Access]}
         dCabinetStatus : DInt := 0;   // Cabinet status (0=OK;1=General power alarm;2=Local power alarm) {x|x|x|x|O}
         dZoneMode : DInt := 4;   // Zone modality (1=Manual;4=Automatic;8=Manual request) {x|x|x|x|O}
         xZoneAlarm : Bool := FALSE;   // Zone alarm {x|x|x|x|O}
         xCalibrationsAllowed : Bool := FALSE;   // Calibration function allowed {x|x|x|x|O}
         dProdModeRequest : DInt := 3;   // Production modality request (1=Out of Production 3= In production) {x|x|x|x|O}
         dProdModeActual : DInt := 3;   // Production modality actual (1=Out of production 3=In production 8=Out of production request 9=In production request) {x|x|x|x|O}
         rgdHeadsActualStatus : Array[0.."CONST_dNumberOfHeadsCycle"] of DInt;   // Head status {x|x|x|x|O}
         tManCmd : Struct
            xSpare : Bool := FALSE;
         END_STRUCT;
      END_STRUCT;
      tHMW : Struct   // {[Unit][Scada unit][Low limit][High limit][Access]}
         xFaultsReset : Bool := FALSE;   // Reset faults {x|x|x|x|O}
         xAutoModeReq : Bool := FALSE;   // Automatic mode request {x|x|x|x|O}
         xManModeReq : Bool := FALSE;   // Manual mode request {x|x|x|x|O}
         xOutOfProdReq : Bool := FALSE;   // Bridge out of production request {x|x|x|x|O}
         xInProdReq : Bool := FALSE;   // Bridge in production request {x|x|x|x|O}
         xGeneralReset : Bool := FALSE;   // General reset {x|x|x|x|M}
         xCutOnBreakEnabled : Bool := FALSE;   // Cut during glass break {x|x|x|x|O}
         xMotorsAndCardsInitialize : Bool := FALSE;   // Motors and cards initialize {x|x|x|x|M}
         dNumberOfLites : DInt := 1;   // Calibration. number of lite on calibration {x|x|1|8|M}
         rgdHeadSelected : Array[0.."CONST_dNumberOfHeadsCycle"] of DInt;   // Calibration. head number selected Cut#x{x|x|1|11|M}
         rgdCutWidthTeo_cmm : Array[0.."CONST_dNumberOfHeadsCycle"] of DInt;   // Calibration. cut width Lite #x theorical [mm/100] {mm/100|mm|200|4000|M}
         rgdCutWidthReal_cmm : Array[0.."CONST_dNumberOfHeadsCycle"] of DInt;   // Calibration. cut width real Lite #x [mm/100] {mm/100|mm|200|4000|M}
         xPositionCalibrationRequest : Bool := FALSE;   // Position calibration request {x|x|x|x|M}
         xForceHeadsHoming : Bool := FALSE;   // Force the homing of the heads {x|x|x|x|M}
         xBridgeOffsetCalibrationRequest : Bool := FALSE;   // Bridge offset calibration request {x|x|x|x|M}
         dMoveBridgeOffset_cmm : DInt := 0;   // Calibration. Move all the heads of this offset {mm/100|mm|-100|100|M}
         dPressureScalerOnSample_perc : DInt := 100;   // Pressure scaler during sample plate [%] {%|%|0|100|O}
         rgxHeadEnabled : Array[0.."CONST_dNumberOfHeadsCycle"] of Bool;   // Head enabled/disabled {x|x|x|x|O}
         tManCmd : Struct
            xBrakeEngage : Bool := FALSE;   // Brake engage all heads {x|x|x|x|O}
            xBrakeRelease : Bool := FALSE;   // Brake release all heads {x|x|x|x|O}
         END_STRUCT;
      END_STRUCT;
   END_VAR
BEGIN
   tHMR.rgdHeadsActualStatus[0] := 3;   // Head #x prod. status (1=Out of production 3=In production 8=Out of production request 9=In production request) {x|x|x|x|O}
   tHMR.rgdHeadsActualStatus[1] := 3;   // Head #x prod. status (1=Out of production 3=In production 8=Out of production request 9=In production request) {x|x|x|x|O}
   tHMR.rgdHeadsActualStatus[2] := 3;   // Head #x prod. status (1=Out of production 3=In production 8=Out of production request 9=In production request) {x|x|x|x|O}
   tHMR.rgdHeadsActualStatus[3] := 3;   // Head #x prod. status (1=Out of production 3=In production 8=Out of production request 9=In production request) {x|x|x|x|O}
   tHMW.rgxHeadEnabled[0] := TRUE;   // Head enabled/disabled {x|x|x|x|O}
   tHMW.rgxHeadEnabled[1] := TRUE;   // Head enabled/disabled {x|x|x|x|O}
   tHMW.rgxHeadEnabled[2] := TRUE;   // Head enabled/disabled {x|x|x|x|O}
   tHMW.rgxHeadEnabled[3] := TRUE;   // Head enabled/disabled {x|x|x|x|O}
   // tHMR.rgdHeadsActualStatus[4] : Head #x prod. status (1=Out of production 3=In production 8=Out of production request 9=In production request) {x|x|x|x|O}
   // tHMW.rgdHeadSelected[0] : Calibration. head number selected Cut#x{x|x|1|11|M}
   // tHMW.rgdHeadSelected[1] : Calibration. head number selected Cut#x{x|x|1|11|M}
   // tHMW.rgdHeadSelected[2] : Calibration. head number selected Cut#x{x|x|1|11|M}
   // tHMW.rgdHeadSelected[3] : Calibration. head number selected Cut#x{x|x|1|11|M}
   // tHMW.rgdHeadSelected[4] : Calibration. head number selected Cut#x{x|x|1|11|M}
   // tHMW.rgdCutWidthTeo_cmm[0] : Calibration. cut width Lite #x theorical [mm/100] {mm/100|mm|200|4000|M}
   // tHMW.rgdCutWidthTeo_cmm[1] : Calibration. cut width Lite #x theorical [mm/100] {mm/100|mm|200|4000|M}
   // tHMW.rgdCutWidthTeo_cmm[2] : Calibration. cut width Lite #x theorical [mm/100] {mm/100|mm|200|4000|M}
   // tHMW.rgdCutWidthTeo_cmm[3] : Calibration. cut width Lite #x theorical [mm/100] {mm/100|mm|200|4000|M}
   // tHMW.rgdCutWidthTeo_cmm[4] : Calibration. cut width Lite #x theorical [mm/100] {mm/100|mm|200|4000|M}
   // tHMW.rgdCutWidthReal_cmm[0] : Calibration. cut width real Lite #x [mm/100] {mm/100|mm|200|4000|M}
   // tHMW.rgdCutWidthReal_cmm[1] : Calibration. cut width real Lite #x [mm/100] {mm/100|mm|200|4000|M}
   // tHMW.rgdCutWidthReal_cmm[2] : Calibration. cut width real Lite #x [mm/100] {mm/100|mm|200|4000|M}
   // tHMW.rgdCutWidthReal_cmm[3] : Calibration. cut width real Lite #x [mm/100] {mm/100|mm|200|4000|M}
   // tHMW.rgdCutWidthReal_cmm[4] : Calibration. cut width real Lite #x [mm/100] {mm/100|mm|200|4000|M}
   // tHMW.rgxHeadEnabled[4] : Head enabled/disabled {x|x|x|x|O}
END_DATA_BLOCK

DATA_BLOCK "Encoder"   // DB17
{ S7_Optimized_Access := 'TRUE' }
VERSION : 0.1
   VAR
      ST_xSystemReset : Bool;   // Reset the system
      ST_xMachineSyncronized : Bool;   // Machine is syncronized
      ST_xMeterPulseArrived : Bool;   // Meter pulse arrived
      OS_xError_YCutMeterGapOutsideLimits : Bool;   // Error. YCut meter gap outside the limits
      OS_xError_MainLineMeterGapOutisdeLimits : Bool;   // Error. Main line meter gap outside the limits
      OS_xError_TimeoutReceivingMeterSignal : Bool;   // Error.Timeout receiving meter signal from main line
      OS_xError_TimeoutReceivingSyncroValue : Bool;   // Error.Timeout receiving syncro value from mainline
      OS_xError_UnexpectedSyncroPulse : Bool;   // Error.Unexpected syncro pulse
      OS_xError_UnexpectedSyncroMessage : Bool;   // Error.Unexpected syncro message
      OSR_xMeterPulse : Bool;   // OSR Meter pulse
      OS_xMeterPulse : Bool;   // OS Meter pulse
      PH_WaitFirstMeter : Bool;   // Waiting first meter pulse
      PH_EndWaitFirstMeter : Bool;   // End waiting first meter pulse
      PH_WaitFirstMeterDataFromMain : Bool;   // Waiting first meter data from main
      PH_EndWaitFirstMeterDataFromMain : Bool;   // End waiting first meter data from main
      PH_WaitMeterPulse : Bool;   // Waiting meter pulse
      PH_EndWaitMeterPulse : Bool;   // End waiting meter pulse
      PH_WaitMeterDataFromMain : Bool;   // Wait meter data from main line
      PH_EndWaitMeterDataFromMain : Bool;   // End wait meter data from main line
      AUX_dActualEncoderValue_cmm : DInt;   // Actual encoder pulse value [mm/100]
      AUX_dActualSpeedValue_cmm_min : DInt;   // Actual lehr speed [cmm/min]
      AUX_dActualSpeedValue_cmm_s : DInt;   // Actual lehr speed [cmm/s]
      AUX_rActualSpeedValue_cmm_ms : Real;   // Actual lehr speed [mm/100 /ms]
      AUX_xNewSyncroReceived : Bool;   // New syncro received from master
      AUX_dNewSyncroValue_cmm : DInt;   // New value of syncro received [mm/100]
      AUX_dLastMainLineValue_cmm : DInt;   // Last main line value syncro [mm/100]
      AUX_dLastStoredSyncroValue_cmm : DInt;   // Last stored syncro value [mm/100]
      AUX_dSyncroGapMainLine_cmm : DInt;   // Syncro gap beetween main line and ycut [mm/100]
      AUX_dMissingSyncroCounter : DInt;   // Missing syncro counter
      AUX_dMeterPulseValue_count : DInt;   // Meter pulse value
      INPUT_dEncoderCounter_count : DInt;   // Encoder counter [count]
      INPUT_dFrequencyCounter_Hz : DInt;   // Frequency counter [Hz]
      INPUT_xMeterPulseArrived : Bool;   // Meter pulse arrived
      INPUT_dMeterPulseValue_count : DInt;   // Meter pulse value [count]
      INPUT_xResetEventAcknowledge : Bool;   // Reset event bit active
      OUTPUT_xCounterEnable : Bool;   // Enable card counter
      OUTPUT_xCounterReset : Bool;   // Card counter reset
      OUTPUT_xResetMeterPulse : Bool;   // Reset meter pulse
      AUX_tmOFFResetMeter : IEC_TIMER;   // Retain meter pulse
      AUX_tmOFFRetainCardReset : IEC_TIMER;   // Retain encoder card reset
   END_VAR
BEGIN
END_DATA_BLOCK

DATA_BLOCK "M256_Manag_Init"   // DB20
{ S7_Optimized_Access := 'TRUE' }
VERSION : 0.1
// stored: InstanceOfName M256_Manager
"M256_Manager"
BEGIN
END_DATA_BLOCK

// folder: 07_ArrayScada

